// TIA Portal project "RRI" (V15.1) (continued)
   PartManagmenent.PartRecept.NazivniPodatki.CILINDRI.MOTOR4[19] := FALSE;
   PartManagmenent.PartRecept.NazivniPodatki.CILINDRI.MOTOR4[20] := FALSE;
   PartManagmenent.PartRecept.NazivniPodatki.CILINDRI.MOTOR5[1] := FALSE;
   PartManagmenent.PartRecept.NazivniPodatki.CILINDRI.MOTOR5[2] := FALSE;
   PartManagmenent.PartRecept.NazivniPodatki.CILINDRI.MOTOR5[3] := FALSE;
   PartManagmenent.PartRecept.NazivniPodatki.CILINDRI.MOTOR5[4] := FALSE;
   PartManagmenent.PartRecept.NazivniPodatki.CILINDRI.MOTOR5[5] := FALSE;
   PartManagmenent.PartRecept.NazivniPodatki.CILINDRI.MOTOR5[6] := FALSE;
   PartManagmenent.PartRecept.NazivniPodatki.CILINDRI.MOTOR5[7] := FALSE;
   PartManagmenent.PartRecept.NazivniPodatki.CILINDRI.MOTOR5[8] := FALSE;
   PartManagmenent.PartRecept.NazivniPodatki.CILINDRI.MOTOR5[9] := FALSE;
   PartManagmenent.PartRecept.NazivniPodatki.CILINDRI.MOTOR5[10] := FALSE;
   PartManagmenent.PartRecept.NazivniPodatki.CILINDRI.MOTOR5[11] := FALSE;
   PartManagmenent.PartRecept.NazivniPodatki.CILINDRI.MOTOR5[12] := FALSE;
   PartManagmenent.PartRecept.NazivniPodatki.CILINDRI.MOTOR5[13] := FALSE;
   PartManagmenent.PartRecept.NazivniPodatki.CILINDRI.MOTOR5[14] := FALSE;
   PartManagmenent.PartRecept.NazivniPodatki.CILINDRI.MOTOR5[15] := FALSE;
   PartManagmenent.PartRecept.NazivniPodatki.CILINDRI.MOTOR5[16] := FALSE;
   PartManagmenent.PartRecept.NazivniPodatki.CILINDRI.MOTOR5[17] := FALSE;
   PartManagmenent.PartRecept.NazivniPodatki.CILINDRI.MOTOR5[18] := FALSE;
   PartManagmenent.PartRecept.NazivniPodatki.CILINDRI.MOTOR5[19] := FALSE;
   PartManagmenent.PartRecept.NazivniPodatki.CILINDRI.MOTOR5[20] := FALSE;
   PartManagmenent.PartRecept.NazivniPodatki.CILINDRI.MOTOR6[1] := FALSE;
   PartManagmenent.PartRecept.NazivniPodatki.CILINDRI.MOTOR6[2] := FALSE;
   PartManagmenent.PartRecept.NazivniPodatki.CILINDRI.MOTOR6[3] := FALSE;
   PartManagmenent.PartRecept.NazivniPodatki.CILINDRI.MOTOR6[4] := FALSE;
   PartManagmenent.PartRecept.NazivniPodatki.CILINDRI.MOTOR6[5] := FALSE;
   PartManagmenent.PartRecept.NazivniPodatki.CILINDRI.MOTOR6[6] := FALSE;
   PartManagmenent.PartRecept.NazivniPodatki.CILINDRI.MOTOR6[7] := FALSE;
   PartManagmenent.PartRecept.NazivniPodatki.CILINDRI.MOTOR6[8] := FALSE;
   PartManagmenent.PartRecept.NazivniPodatki.CILINDRI.MOTOR6[9] := FALSE;
   PartManagmenent.PartRecept.NazivniPodatki.CILINDRI.MOTOR6[10] := FALSE;
   PartManagmenent.PartRecept.NazivniPodatki.CILINDRI.MOTOR6[11] := FALSE;
   PartManagmenent.PartRecept.NazivniPodatki.CILINDRI.MOTOR6[12] := FALSE;
   PartManagmenent.PartRecept.NazivniPodatki.CILINDRI.MOTOR6[13] := FALSE;
   PartManagmenent.PartRecept.NazivniPodatki.CILINDRI.MOTOR6[14] := FALSE;
   PartManagmenent.PartRecept.NazivniPodatki.CILINDRI.MOTOR6[15] := FALSE;
   PartManagmenent.PartRecept.NazivniPodatki.CILINDRI.MOTOR6[16] := FALSE;
   PartManagmenent.PartRecept.NazivniPodatki.CILINDRI.MOTOR6[17] := FALSE;
   PartManagmenent.PartRecept.NazivniPodatki.CILINDRI.MOTOR6[18] := FALSE;
   PartManagmenent.PartRecept.NazivniPodatki.CILINDRI.MOTOR6[19] := FALSE;
   PartManagmenent.PartRecept.NazivniPodatki.CILINDRI.MOTOR6[20] := FALSE;
   PartManagmenent.PartRecept.TrenutniPodatki.trenutni_pomik := 0;
   PartManagmenent.PartRecept.Oblika.s1[0] := FALSE;
   PartManagmenent.PartRecept.Oblika.s1[1] := FALSE;
   PartManagmenent.PartRecept.Oblika.s1[2] := FALSE;
   PartManagmenent.PartRecept.Oblika.s1[3] := FALSE;
   PartManagmenent.PartRecept.Oblika.s1[4] := FALSE;
   PartManagmenent.PartRecept.Oblika.s1[5] := FALSE;
   PartManagmenent.PartRecept.Oblika.s1[6] := FALSE;
   PartManagmenent.PartRecept.Oblika.s1[7] := FALSE;
   PartManagmenent.PartRecept.Oblika.s1[8] := FALSE;
   PartManagmenent.PartRecept.Oblika.s1[9] := FALSE;
   PartManagmenent.PartRecept.Oblika.s1[10] := FALSE;
   PartManagmenent.PartRecept.Oblika.s1[11] := FALSE;
   PartManagmenent.PartRecept.Oblika.s1[12] := FALSE;
   PartManagmenent.PartRecept.Oblika.s1[13] := FALSE;
   PartManagmenent.PartRecept.Oblika.s1[14] := FALSE;
   PartManagmenent.PartRecept.Oblika.s1[15] := FALSE;
   PartManagmenent.PartRecept.Oblika.s1[16] := FALSE;
   PartManagmenent.PartRecept.Oblika.s1[17] := FALSE;
   PartManagmenent.PartRecept.Oblika.s1[18] := FALSE;
   PartManagmenent.PartRecept.Oblika.s1[19] := FALSE;
   PartManagmenent.PartRecept.Oblika.s1[20] := FALSE;
   PartManagmenent.PartRecept.Oblika.s2[0] := FALSE;
   PartManagmenent.PartRecept.Oblika.s2[1] := FALSE;
   PartManagmenent.PartRecept.Oblika.s2[2] := FALSE;
   PartManagmenent.PartRecept.Oblika.s2[3] := FALSE;
   PartManagmenent.PartRecept.Oblika.s2[4] := FALSE;
   PartManagmenent.PartRecept.Oblika.s2[5] := FALSE;
   PartManagmenent.PartRecept.Oblika.s2[6] := FALSE;
   PartManagmenent.PartRecept.Oblika.s2[7] := FALSE;
   PartManagmenent.PartRecept.Oblika.s2[8] := FALSE;
   PartManagmenent.PartRecept.Oblika.s2[9] := FALSE;
   PartManagmenent.PartRecept.Oblika.s2[10] := FALSE;
   PartManagmenent.PartRecept.Oblika.s2[11] := FALSE;
   PartManagmenent.PartRecept.Oblika.s2[12] := FALSE;
   PartManagmenent.PartRecept.Oblika.s2[13] := FALSE;
   PartManagmenent.PartRecept.Oblika.s2[14] := FALSE;
   PartManagmenent.PartRecept.Oblika.s2[15] := FALSE;
   PartManagmenent.PartRecept.Oblika.s2[16] := FALSE;
   PartManagmenent.PartRecept.Oblika.s2[17] := FALSE;
   PartManagmenent.PartRecept.Oblika.s2[18] := FALSE;
   PartManagmenent.PartRecept.Oblika.s2[19] := FALSE;
   PartManagmenent.PartRecept.Oblika.s2[20] := FALSE;
   PartManagmenent.xMerkers[0] := FALSE;
   PartManagmenent.xMerkers[1] := FALSE;
END_DATA_BLOCK

DATA_BLOCK "FB_TcConvert_DB_TC1_ToolTemeprature"   // DB4
{ S7_Optimized_Access := 'TRUE' }
VERSION : 0.1
// stored: InstanceOfName FB_TcConvert
"FB_TcConvert"
BEGIN
END_DATA_BLOCK

DATA_BLOCK "FB_TcConvert_DB_TC2_ToolTemeprature"   // DB5
{ S7_Optimized_Access := 'TRUE' }
VERSION : 0.1
// stored: InstanceOfName FB_TcConvert
"FB_TcConvert"
BEGIN
END_DATA_BLOCK

DATA_BLOCK "FB_AKDstartup_DB_AKD1"   // DB6
{ S7_Optimized_Access := 'TRUE' }
VERSION : 0.1
// stored: InstanceOfName FB_AKDstartup
"FB_AKDstartup"
BEGIN
END_DATA_BLOCK

DATA_BLOCK "FB_AKDstartup_DB_TC4"   // DB7
{ S7_Optimized_Access := 'TRUE' }
VERSION : 0.1
// stored: InstanceOfName FB_AKDstartup
"FB_AKDstartup"
BEGIN
END_DATA_BLOCK

DATA_BLOCK "FB_TcConvert_DB_tc4"   // DB8
{ S7_Optimized_Access := 'TRUE' }
VERSION : 0.1
// stored: InstanceOfName FB_TcConvert
"FB_TcConvert"
BEGIN
END_DATA_BLOCK

DATA_BLOCK "FB_RTDConvert_DB_RTD1"   // DB9
{ S7_Optimized_Access := 'TRUE' }
VERSION : 0.1
// stored: InstanceOfName FB_RTDConvert
"FB_RTDConvert"
BEGIN
END_DATA_BLOCK

DATA_BLOCK "FB_RTDConvert_DB_RTD2"   // DB10
{ S7_Optimized_Access := 'TRUE' }
VERSION : 0.1
// stored: InstanceOfName FB_RTDConvert
"FB_RTDConvert"
BEGIN
END_DATA_BLOCK

DATA_BLOCK "FB_RTDConvert_DB_RTD3"   // DB11
{ S7_Optimized_Access := 'TRUE' }
VERSION : 0.1
// stored: InstanceOfName FB_RTDConvert
"FB_RTDConvert"
BEGIN
END_DATA_BLOCK

DATA_BLOCK "FB_RTDConvert_DB_RTD4"   // DB12
{ S7_Optimized_Access := 'TRUE' }
VERSION : 0.1
// stored: InstanceOfName FB_RTDConvert
"FB_RTDConvert"
BEGIN
END_DATA_BLOCK

DATA_BLOCK "LMqtt_Publisher_DB"   // DB13
{ S7_Optimized_Access := 'TRUE' }
VERSION : 0.1
// stored: InstanceOfName LMqtt_Publisher
"LMqtt_Publisher"
BEGIN
END_DATA_BLOCK

DATA_BLOCK "FB_concatScrings_DB"   // DB18
{ S7_Optimized_Access := 'TRUE' }
VERSION : 0.1
// stored: InstanceOfName FB_concatScrings
"FB_concatScrings"
BEGIN
END_DATA_BLOCK

DATA_BLOCK "DB_rPMCalculator"   // DB19
{ S7_Optimized_Access := 'TRUE' }
VERSION : 0.1
   VAR RETAIN
      Press_one : Struct
         p_trig : Bool;
         iCurrentCounter : Int;
         rCurrentSpeed : Int;
         PulseTimer : TON_TIME;
         xcalculateRPM : Bool;
      END_STRUCT;
   END_VAR
BEGIN
END_DATA_BLOCK

DATA_BLOCK "LMqtt_Publisher_DB1"   // DB22
{ S7_Optimized_Access := 'TRUE' }
VERSION : 0.1
// stored: InstanceOfName LMqtt_Publisher
"LMqtt_Publisher"
BEGIN
END_DATA_BLOCK

DATA_BLOCK "FB_concatScrings_DB1"   // DB23
{ S7_Optimized_Access := 'TRUE' }
VERSION : 0.1
// stored: InstanceOfName FB_concatScrings
"FB_concatScrings"
BEGIN
END_DATA_BLOCK

DATA_BLOCK "FB_CONCAT_STRINGS_FOR_MQTT_DB"   // DB24
{ S7_Optimized_Access := 'TRUE' }
VERSION : 0.1
// stored: InstanceOfName FB_CONCAT_STRINGS_FOR_MQTT
"FB_CONCAT_STRINGS_FOR_MQTT"
BEGIN
END_DATA_BLOCK

DATA_BLOCK "LMqtt_Publisher_1_DB"   // DB25
{ S7_Optimized_Access := 'TRUE' }
VERSION : 0.1
// stored: InstanceOfName LMqtt_Publisher_1
"LMqtt_Publisher_1"
BEGIN
END_DATA_BLOCK

DATA_BLOCK "DB_TESTWSTRING"   // DB26
{ S7_Optimized_Access := 'TRUE' }
VERSION : 0.1
   VAR
      wstring_test : WString[1000];
   END_VAR
BEGIN
END_DATA_BLOCK

DATA_BLOCK "FB_CONCAT_STRINGS_FOR_MQTT_DB_1"   // DB27
{ S7_Optimized_Access := 'TRUE' }
VERSION : 0.1
// stored: InstanceOfName FB_CONCAT_STRINGS_FOR_MQTT
"FB_CONCAT_STRINGS_FOR_MQTT"
BEGIN
END_DATA_BLOCK

DATA_BLOCK "FB_CONCAT_STRINGS_FOR_MQTT_1_DB"   // DB28
{ S7_Optimized_Access := 'TRUE' }
VERSION : 0.1
// stored: InstanceOfName FB_CONCAT_STRINGS_FOR_MQTT_1
"FB_CONCAT_STRINGS_FOR_MQTT_1"
BEGIN
END_DATA_BLOCK

DATA_BLOCK "FB_saveConcat_DB"   // DB29
{ S7_Optimized_Access := 'TRUE' }
VERSION : 0.1
// stored: InstanceOfName FB_saveConcat
"FB_saveConcat"
BEGIN
END_DATA_BLOCK

DATA_BLOCK "FB_AKD_DB_AKD1"   // DB30
{ S7_Optimized_Access := 'TRUE' }
VERSION : 0.1
// stored: InstanceOfName FB_AKD
"FB_AKD"
BEGIN
END_DATA_BLOCK

DATA_BLOCK "_AKD1"   // DB32
{ S7_Optimized_Access := 'TRUE' }
VERSION : 0.1
// stored: InstanceOfName PTC_1000_resistanceCalculation
"PTC_1000_resistanceCalculation"
BEGIN
END_DATA_BLOCK

DATA_BLOCK "FB_EgasiMotorControl_DB_M1"   // DB35
{ S7_Optimized_Access := 'TRUE' }
VERSION : 0.1
// stored: InstanceOfName FB_EgasiMotorControl
"FB_EgasiMotorControl"
BEGIN
END_DATA_BLOCK

DATA_BLOCK "DB_safetyActuator"   // DB36
{ S7_Optimized_Access := 'TRUE' }
VERSION : 0.1
   VAR RETAIN
      On_timer : Array[0..1] of TON_TIME;
      timerOut : Bool;
   END_VAR
BEGIN
END_DATA_BLOCK

DATA_BLOCK "FB_EgasiMotorControl_DB_M2"   // DB37
{ S7_Optimized_Access := 'TRUE' }
VERSION : 0.1
// stored: InstanceOfName FB_EgasiMotorControl
"FB_EgasiMotorControl"
BEGIN
END_DATA_BLOCK

DATA_BLOCK "FB_EgasiMotorControl_DB_M3"   // DB38
{ S7_Optimized_Access := 'TRUE' }
VERSION : 0.1
// stored: InstanceOfName FB_EgasiMotorControl
"FB_EgasiMotorControl"
BEGIN
END_DATA_BLOCK

DATA_BLOCK "FB_EgasiMotorControl_DB_M4"   // DB39
{ S7_Optimized_Access := 'TRUE' }
VERSION : 0.1
// stored: InstanceOfName FB_EgasiMotorControl
"FB_EgasiMotorControl"
BEGIN
END_DATA_BLOCK

DATA_BLOCK "FB_EgasiMotorControl_DB_M5"   // DB40
{ S7_Optimized_Access := 'TRUE' }
VERSION : 0.1
// stored: InstanceOfName FB_EgasiMotorControl
"FB_EgasiMotorControl"
BEGIN
END_DATA_BLOCK

DATA_BLOCK "DB_EGASI_MOTOR_BASE"   // DB41
{ S7_Optimized_Access := 'TRUE' }
VERSION : 0.1
   VAR RETAIN
      MOTOR : Array[1..5] of "EGASI_MOTOR_CONTROL";
   END_VAR
BEGIN
END_DATA_BLOCK

DATA_BLOCK "DB_PARTS_DATABASE"   // DB42
{ S7_Optimized_Access := 'TRUE' }
VERSION : 0.1
BEGIN
END_DATA_BLOCK

DATA_BLOCK "DB_RRI_Izdelki"   // DB43
{ S7_Optimized_Access := 'TRUE' }
VERSION : 0.1
   VAR RETAIN
      "1x2-Cell" : "RRI_izdelki";
      "1x4-Cell" : "RRI_izdelki";
      "1x6-Cell" : "RRI_izdelki";
      "1x8-Cell" : "RRI_izdelki";
      "2x2-Cell" : "RRI_izdelki";
      "2x4-Cell" : "RRI_izdelki";
      "2x6-Cell" : "RRI_izdelki";
      "2x8-Cell" : "RRI_izdelki";
      "39900-8" : "RRI_izdelki";
      "39900-9" : "RRI_izdelki";
   END_VAR
BEGIN
   "1x2-Cell".NazivniPodatki.st_pomikov := 2;
   "1x2-Cell".NazivniPodatki.st_celic := 2;
   "1x2-Cell".NazivniPodatki.st_vrst := 1;
   "1x4-Cell".NazivniPodatki.st_pomikov := 4;
   "1x4-Cell".NazivniPodatki.st_celic := 4;
   "1x4-Cell".NazivniPodatki.st_vrst := 1;
   "1x6-Cell".NazivniPodatki.st_pomikov := 6;
   "1x6-Cell".NazivniPodatki.st_celic := 6;
   "1x6-Cell".NazivniPodatki.st_vrst := 1;
   "1x8-Cell".NazivniPodatki.st_celic := 8;
   "1x8-Cell".NazivniPodatki.st_pomikov := 8;
   "1x8-Cell".NazivniPodatki.st_vrst := 1;
   "2x2-Cell".NazivniPodatki.st_pomikov := 2;
   "2x2-Cell".NazivniPodatki.st_celic := 2;
   "2x2-Cell".NazivniPodatki.st_vrst := 2;
   "2x4-Cell".NazivniPodatki.st_pomikov := 4;
   "2x4-Cell".NazivniPodatki.st_celic := 4;
   "2x4-Cell".NazivniPodatki.st_vrst := 2;
   "2x6-Cell".NazivniPodatki.st_pomikov := 6;
   "2x6-Cell".NazivniPodatki.st_celic := 6;
   "2x6-Cell".NazivniPodatki.st_vrst := 2;
   "2x8-Cell".NazivniPodatki.st_pomikov := 8;
   "2x8-Cell".NazivniPodatki.st_celic := 8;
   "2x8-Cell".NazivniPodatki.st_vrst := 2;
END_DATA_BLOCK

DATA_BLOCK "FB_CYLINDER_CONTROL_DB"   // DB44
{ S7_Optimized_Access := 'TRUE' }
VERSION : 0.1
// stored: InstanceOfName FB_CYLINDER_CONTROL
"FB_CYLINDER_CONTROL"
BEGIN
END_DATA_BLOCK

DATA_BLOCK "FB_VerifyTheFormLerning_DB"   // DB47
{ S7_Optimized_Access := 'TRUE' }
VERSION : 0.1
// stored: InstanceOfName FB_VerifyTheFormLerning
"FB_VerifyTheFormLerning"
BEGIN
END_DATA_BLOCK

DATA_BLOCK "DB_newGlobalDataForChangeParrt"   // DB48
{ S7_Optimized_Access := 'TRUE' }
VERSION : 0.1
   VAR RETAIN
      ud_GlobalFeedCounter : UDInt;
      DATA : "M_position";
      changePartCounter : UDInt;
      strip : Array[0..20] of "STRIP_SEGMENT";
   END_VAR
BEGIN
   DATA.POSITION_INSIDE_TOOL.M1 := 5;
   DATA.POSITION_INSIDE_TOOL.M2 := 8;
   DATA.POSITION_INSIDE_TOOL.M3 := 10;
   DATA.POSITION_INSIDE_TOOL.M4 := 14;
   DATA.POSITION_INSIDE_TOOL.M5 := 17;
   DATA.POSITION_INSIDE_TOOL.TOOL_MAX_FEED := 17;
END_DATA_BLOCK

DATA_BLOCK "FB_CYLINDER_CONTROL_PIPILINE_DB"   // DB49
{ S7_Optimized_Access := 'TRUE' }
VERSION : 0.1
// stored: InstanceOfName FB_CYLINDER_CONTROL_PIPILINE
"FB_CYLINDER_CONTROL_PIPILINE"
BEGIN
END_DATA_BLOCK

// folder: AKD

DATA_BLOCK "DB_AKD"   // DB31
{ S7_Optimized_Access := 'TRUE' }
VERSION : 0.1
BEGIN
END_DATA_BLOCK

// folder: AKD/PNU

DATA_BLOCK "AKD_PNU_DATA"   // DB33
{ S7_Optimized_Access := 'TRUE' }
VERSION : 0.1
   VAR
      AKD1 : Struct
         PNU_DATA : "PNU_DATA";
         PNU_userSETTINGS : Struct
            xRadAKDTemp : Bool;
            xReadAkdTempInC : Bool;
            PNU_const : Struct
               AKD_TEMP : Struct
                  PNU_number : Int := 2257;
                  PNU_subIndex : Int := 0;
                  PNU_type : Word := 16#43;
               END_STRUCT;
               AKD_TEMP_C : Struct
                  PNU_number : Int := 2258;
                  PNU_subIndex : Int := 0;
                  PNU_type : Word := 16#43;
               END_STRUCT;
            END_STRUCT;
         END_STRUCT;
      END_STRUCT;
   END_VAR
BEGIN
END_DATA_BLOCK

DATA_BLOCK "AKD1_PNU"   // DB34
{ S7_Optimized_Access := 'FALSE' }
AUTHOR : jcoleman
FAMILY : PNU
VERSION : 2.0
// stored: InstanceOfName AKD_PNU_v02
"AKD_PNU_v02"
BEGIN
END_DATA_BLOCK

// folder: MQTT

DATA_BLOCK "LMqtt_Status"   // DB14
{ S7_Optimized_Access := 'TRUE' }
VERSION : 0.1
   VAR
      mqtt_1 : Struct
         xtcpEsablished : Bool;   // True if the TCP connection has been
         xmqttEstavlished : Bool;   // True if the MQTT connection has been established
         xpublished : Bool;   // True, if the message has arrived successfully at
         xbusy : Bool;   // True, while a message or ping is sent to the
         xerror : Bool;   // True if there is an error
         istatusID : Int;   // State that cause the error
         status : DWord;   // Error message
      END_STRUCT;
   END_VAR
BEGIN
END_DATA_BLOCK

DATA_BLOCK "instPublisherDB"   // DB15
{ S7_Optimized_Access := 'TRUE' }
VERSION : 0.1
// stored: InstanceOfName LMqtt_Publisher
"LMqtt_Publisher"
BEGIN
END_DATA_BLOCK

DATA_BLOCK "LMqtt_Data"   // DB16
{ S7_Optimized_Access := 'TRUE' }
VERSION : 0.1
   VAR
      dataTcp : "typeTcpConnParam";
      dataMqtt : "typeMqttParam";
   END_VAR
BEGIN
   dataMqtt.connectFlag.cleanSession := 1;
   dataMqtt.connectFlag.will := 0;
   dataMqtt.connectFlag.willQoS_1 := 0;
   dataMqtt.connectFlag.willRetain := 0;
   dataMqtt.clientIdentifier := 'S7-1200-PLC';
   dataMqtt.willTopic := '/final';
   dataMqtt.willMessage := 'Das wars';
   dataTcp.hwIdentifier := 64;
   dataTcp.connectionID := 16#2;
   dataTcp.ipAdressBroker[0] := 192;
   dataMqtt.topic := 'data/s71200';
   dataMqtt.message := 'My first message';
   dataMqtt.publishFlag.qualityOfService := 1;
   dataMqtt.keepAlive := 0;
   dataTcp.localPort := 2000;
   dataTcp.mqttPort := 1883;
   dataMqtt.connectFlag.password := 0;
   dataMqtt.connectFlag.userName := 0;
   dataMqtt.userName := 'simatic';
   dataMqtt.password := 'Anna';
   dataTcp.ipAdressBroker[1] := 168;
   dataTcp.ipAdressBroker[2] := 1;
   dataTcp.ipAdressBroker[3] := 1;
END_DATA_BLOCK

DATA_BLOCK "LMqtt_publish"   // DB17
{ S7_Optimized_Access := 'TRUE' }
VERSION : 0.1
   VAR
      LMqtt : Struct
         xenable : Bool;
         epublish : Bool;
         sStringToPublish : String;
      END_STRUCT;
      randomstrinmg : String;
   END_VAR
BEGIN
END_DATA_BLOCK

// folder: MQTT/userData

DATA_BLOCK "MQTT_DB"   // DB21
{ S7_Optimized_Access := 'TRUE' }
VERSION : 0.1
   VAR RETAIN
      MQTT_CLIEENTS : Array[0..1] of "typeMqttData";
   END_VAR
   VAR
      MQTT_CLIENTS_WSTRING : Array[0..1] of "typeMqttData_1";
   END_VAR
BEGIN
   MQTT_CLIEENTS[0].mqttTcpParam.hwIdentifier := 64;
   MQTT_CLIEENTS[0].mqttTcpParam.connectionID := 16#0003;
   MQTT_CLIEENTS[0].mqttTcpParam.ipAdressBroker[0] := 16#C0;
   MQTT_CLIEENTS[0].mqttTcpParam.ipAdressBroker[1] := 16#A8;
   MQTT_CLIEENTS[0].mqttTcpParam.ipAdressBroker[2] := 16#01;
   MQTT_CLIEENTS[0].mqttTcpParam.ipAdressBroker[3] := 16#01;
   MQTT_CLIEENTS[0].mqttTcpParam.localPort := 2001;
   MQTT_CLIEENTS[0].mqttTcpParam.mqttPort := 1883;
   MQTT_CLIEENTS[0].mqttParam.connectFlag.cleanSession := TRUE;
   MQTT_CLIEENTS[0].mqttParam.clientIdentifier := 'S7-1200-PLC2';
   MQTT_CLIEENTS[0].mqttParam.willTopic := '/final2';
   MQTT_CLIEENTS[0].mqttParam.topic := 'data/s71200/RTDvalues';
   MQTT_CLIEENTS[0].mqttParam.message := '{"temperature1":                  -1.0000,"temperature2":                  -1.0000,"temperature3":                  22.8000,"temperature4":                  -1.0000}';
   MQTT_CLIEENTS[0].mqttParam.connectFlag.will := FALSE;
   MQTT_CLIEENTS[0].mqttParam.connectFlag.willQoS_1 := FALSE;
   MQTT_CLIEENTS[0].mqttParam.connectFlag.willQoS_2 := FALSE;
   MQTT_CLIEENTS[0].mqttParam.connectFlag.willRetain := FALSE;
   MQTT_CLIEENTS[0].mqttParam.connectFlag.password := FALSE;
   MQTT_CLIEENTS[0].mqttParam.connectFlag.userName := FALSE;
   MQTT_CLIEENTS[0].mqttParam.publishFlag.qualityOfService := 0;
   MQTT_CLIEENTS[0].mqttParam.publishFlag.retain := FALSE;
   MQTT_CLIEENTS[0].mqttParam.keepAlive := 16#000A;
   MQTT_CLIEENTS[0].mqttParam.packetIdentifier := 16#0010;
   MQTT_CLIEENTS[0].mqttParam.willMessage := 'das';
   MQTT_CLIEENTS[0].mqttParam.userName := 'Simatic';
   MQTT_CLIEENTS[0].mqttParam.password := 'Anna';
   MQTT_CLIEENTS[0].mqttUserControl.xEnable := TRUE;
   MQTT_CLIEENTS[0].mqttUserControl.xPusblish := FALSE;
   MQTT_CLIEENTS[0].mqttUserControl.sStringToPublish := '{"temperature1":                  -1.0000,"temperature2":                  -1.0000,"temperature3":                  22.8000,"temperature4":                  -1.0000}';
   MQTT_CLIEENTS[0].mqttUserControl.Status.xtcpEsablished := TRUE;
   MQTT_CLIEENTS[0].mqttUserControl.Status.xmqttEstavlished := TRUE;
   MQTT_CLIEENTS[0].mqttUserControl.Status.xpublished := FALSE;
   MQTT_CLIEENTS[0].mqttUserControl.Status.xbusy := FALSE;
   MQTT_CLIEENTS[0].mqttUserControl.Status.xerror := FALSE;
   MQTT_CLIEENTS[0].mqttUserControl.Status.istatusID := 0;
   MQTT_CLIEENTS[0].mqttUserControl.Status.status := 16#0000_0000;
   MQTT_CLIEENTS[1].mqttTcpParam.hwIdentifier := 0;
   MQTT_CLIEENTS[1].mqttTcpParam.connectionID := 16#0000;
   MQTT_CLIEENTS[1].mqttTcpParam.ipAdressBroker[0] := 16#00;
   MQTT_CLIEENTS[1].mqttTcpParam.ipAdressBroker[1] := 16#00;
   MQTT_CLIEENTS[1].mqttTcpParam.ipAdressBroker[2] := 16#00;
   MQTT_CLIEENTS[1].mqttTcpParam.ipAdressBroker[3] := 16#00;
   MQTT_CLIEENTS[1].mqttTcpParam.localPort := 0;
   MQTT_CLIEENTS[1].mqttTcpParam.mqttPort := 0;
   MQTT_CLIEENTS[1].mqttParam.connectFlag.cleanSession := FALSE;
   MQTT_CLIEENTS[1].mqttParam.connectFlag.will := FALSE;
   MQTT_CLIEENTS[1].mqttParam.connectFlag.willQoS_1 := FALSE;
   MQTT_CLIEENTS[1].mqttParam.connectFlag.willQoS_2 := FALSE;
   MQTT_CLIEENTS[1].mqttParam.connectFlag.willRetain := FALSE;
   MQTT_CLIEENTS[1].mqttParam.connectFlag.password := FALSE;
   MQTT_CLIEENTS[1].mqttParam.connectFlag.userName := FALSE;
   MQTT_CLIEENTS[1].mqttParam.publishFlag.qualityOfService := 0;
   MQTT_CLIEENTS[1].mqttParam.publishFlag.retain := FALSE;
   MQTT_CLIEENTS[1].mqttParam.keepAlive := 16#000A;
   MQTT_CLIEENTS[1].mqttParam.packetIdentifier := 16#0010;
   MQTT_CLIEENTS[1].mqttParam.clientIdentifier := '';
   MQTT_CLIEENTS[1].mqttParam.willTopic := '';
   MQTT_CLIEENTS[1].mqttParam.willMessage := '';
   MQTT_CLIEENTS[1].mqttParam.userName := '';
   MQTT_CLIEENTS[1].mqttParam.password := '';
   MQTT_CLIEENTS[1].mqttParam.topic := '';
   MQTT_CLIEENTS[1].mqttParam.message := '';
   MQTT_CLIEENTS[1].mqttUserControl.xEnable := FALSE;
   MQTT_CLIEENTS[1].mqttUserControl.xPusblish := FALSE;
   MQTT_CLIEENTS[1].mqttUserControl.sStringToPublish := '';
   MQTT_CLIEENTS[1].mqttUserControl.Status.xtcpEsablished := FALSE;
   MQTT_CLIEENTS[1].mqttUserControl.Status.xmqttEstavlished := FALSE;
   MQTT_CLIEENTS[1].mqttUserControl.Status.xpublished := FALSE;
   MQTT_CLIEENTS[1].mqttUserControl.Status.xbusy := FALSE;
   MQTT_CLIEENTS[1].mqttUserControl.Status.xerror := FALSE;
   MQTT_CLIEENTS[1].mqttUserControl.Status.istatusID := 0;
   MQTT_CLIEENTS[1].mqttUserControl.Status.status := 16#0000_0000;
   MQTT_CLIENTS_WSTRING[0].mqttParam.topic := 'data/s71200/testValues';
   MQTT_CLIENTS_WSTRING[0].mqttParam.password := 'Anna';
   MQTT_CLIENTS_WSTRING[0].mqttParam.userName := 'Simatic';
   MQTT_CLIENTS_WSTRING[0].mqttParam.willMessage := 'das';
   MQTT_CLIENTS_WSTRING[0].mqttParam.willTopic := '/final2';
   MQTT_CLIENTS_WSTRING[0].mqttParam.clientIdentifier := 'S7-1200-WS';
   MQTT_CLIENTS_WSTRING[0].mqttParam.packetIdentifier := 16#0010;
   MQTT_CLIENTS_WSTRING[0].mqttParam.keepAlive := 16#000A;
   MQTT_CLIENTS_WSTRING[0].mqttParam.connectFlag.cleanSession := TRUE;
   MQTT_CLIENTS_WSTRING[0].mqttTcpParam.mqttPort := 1883;
   MQTT_CLIENTS_WSTRING[0].mqttTcpParam.localPort := 2003;
   MQTT_CLIENTS_WSTRING[0].mqttTcpParam.ipAdressBroker[3] := 16#01;
   MQTT_CLIENTS_WSTRING[0].mqttTcpParam.ipAdressBroker[2] := 16#01;
   MQTT_CLIENTS_WSTRING[0].mqttTcpParam.ipAdressBroker[1] := 16#A8;
   MQTT_CLIENTS_WSTRING[0].mqttTcpParam.ipAdressBroker[0] := 16#C0;
   MQTT_CLIENTS_WSTRING[0].mqttTcpParam.connectionID := 16#0006;
   MQTT_CLIENTS_WSTRING[0].mqttTcpParam.hwIdentifier := 64;
END_DATA_BLOCK

// folder: NodeRed

DATA_BLOCK "DB_DATAFORCOMMUNICATION"   // DB1
{ S7_Optimized_Access := 'FALSE' }
VERSION : 0.1
   VAR
      rTC1_ToolTemperature1 : Real;
      rTC2_ToolTemeprature2 : Real;
      rTC3_TempEnvierment : Real;
      rTC4_Temp : Real;
      iPresaHitrost : Int;
      uPresaStevec : UDInt;
      xPresaON : Int;
      r_RTD_c0 : Real;   // temp ohišja aktuatorja
      r_RTD_c1 : Real;   // ohišje orodja
      r_RTD_c2 : Real;
      r_RTD_c3 : Real;
      r_ActuatorMaxForce : Real;
      r_ActuatorMinForce : Real;
      r_EgasiTemperaturaAktuatorja : Real;
      r_M1_temperature : Real;
      r_M2_temperature : Real;
      r_M3_temperature : Real;
      r_M4_temperature : Real;
      r_M5_temperature : Real;
      r_M1_MaxForce : Real;
      r_M2_MaxForce : Real;
      r_M3_MaxForce : Real;
      r_M4_MaxForce : Real;
      r_M5_MaxForce : Real;
      i_StevecPomika : Int;
      test : Int;
      iHMIpartNumber : Int;   // Part number -> Manual
      iHmiLastPartNumber : Int;
      iOperationMode : Int;   // 0 -> MANUAL 1->AUTO
   END_VAR
BEGIN
END_DATA_BLOCK

DATA_BLOCK "DB_MotorData"   // DB45
{ S7_Optimized_Access := 'FALSE' }
VERSION : 0.1
   VAR
      M1_status : "UDT_MotorDataStatus";
      M2_status : "UDT_MotorDataStatus";
      M3_status : "UDT_MotorDataStatus";
      M4_status : "UDT_MotorDataStatus";
      M5_status : "UDT_MotorDataStatus";
   END_VAR
BEGIN
END_DATA_BLOCK

DATA_BLOCK "DB_MotorControl"   // DB46
{ S7_Optimized_Access := 'FALSE' }
VERSION : 0.1
   VAR
      HMI_M1 : "UDT_MotorControl";
      HMI_M2 : "UDT_MotorControl";
      HMI_M3 : "UDT_MotorControl";
      HMI_M4 : "UDT_MotorControl";
      HMI_M5 : "UDT_MotorControl";
      xOverRideControl : Bool;   // 1 - HMI, 0 - PLC - MOTOR STATUS , CONTRO mode HMI
      xManualMode : Bool;
      xDEMO_or_AutomaticMode : Bool;   // 0 - automatic, 1- demo
      xHMI_resetPomikna0 : Bool;
      xHMI_Manual_or_automatic_production : Bool;   // 1-MANUAL, 0-AUTOMATIC - prodution
      DTL_forProductionID : DTL;
      Static_1 : UDInt;
   END_VAR
BEGIN
END_DATA_BLOCK

// folder: System blocks/Program resources

DATA_BLOCK "xPresaOFF"   // DB20
{ S7_Optimized_Access := 'TRUE' }
AUTHOR : Simatic
FAMILY : IEC
NAME : IEC_TMR
VERSION : 1.0
// stored: InstanceOfName IEC_TIMER
"IEC_TIMER"
BEGIN
END_DATA_BLOCK

// folder: (top level)

FUNCTION_BLOCK "FB_TcConvert"   // FB1, LAD
{ S7_Optimized_Access := 'TRUE' }
VERSION : 0.1
// Convert Thermocoupler input to the °C value
   VAR_INPUT
      i_wTC_value : Word;
      i_rCalibrationFactor : Real;
   END_VAR
   VAR_OUTPUT
      q_rTemperature : Real;
   END_VAR
   VAR RETAIN
      _rConvertedValue : Real;
   END_VAR
BEGIN

REGION Network 2 (SCL)

   //Input value 254 (DEC) = 25.5°C
   //32767 - overflow or error
   IF #i_wTC_value = 32767 THEN
       #q_rTemperature := -1.0;
       RETURN;
   END_IF;

   #q_rTemperature := WORD_TO_DINT( #i_wTC_value) / 10.0-#i_rCalibrationFactor;
END_REGION
END_FUNCTION_BLOCK

FUNCTION_BLOCK "FB_AKDstartup"   // FB2, LAD
{ S7_Optimized_Access := 'TRUE' }
VERSION : 0.1
   VAR_INPUT
      i_xFaultFeedback : Bool;   // AKD drive fault - open (0) if error
      i_xStart : Bool;   // Run startup Sequence
   END_VAR
   VAR_OUTPUT
      q_xHwEnable : Bool;
      q_xSTOEnable : Bool;
      q_xAKDPower : Bool;
      q_xSoftwareEnable : Bool;
   END_VAR
   VAR
      TON_TIMER : Array[0..1] of TON_TIME;
      TOFF_TIMER : Array[0..1] of TOF_TIME;
   END_VAR
BEGIN

REGION Network 1
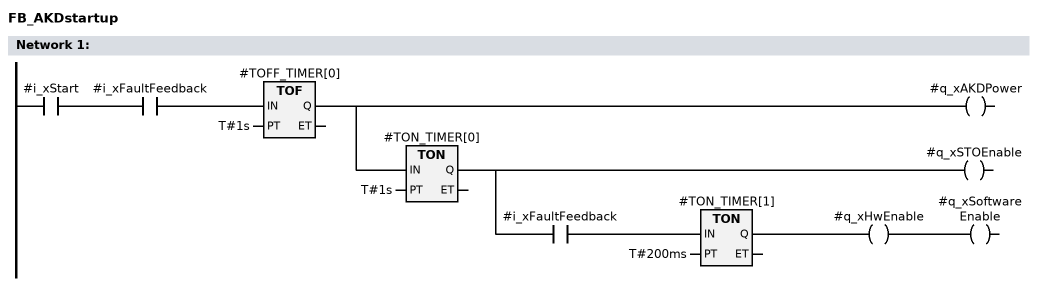
   #TOFF_TIMER[0].TOF(IN := #i_xStart AND #i_xFaultFeedback, PT := T#1s);
   #q_xAKDPower := #TOFF_TIMER[0].Q;
   #TON_TIMER[0].TON(IN := #TOFF_TIMER[0].Q, PT := T#1s);
   #q_xSTOEnable := #TON_TIMER[0].Q;
   #TON_TIMER[1].TON(IN := #TON_TIMER[0].Q AND #i_xFaultFeedback, PT := T#200ms);
   #q_xHwEnable := #TON_TIMER[1].Q;
   #q_xSoftwareEnable := #TON_TIMER[1].Q;
END_REGION
END_FUNCTION_BLOCK

FUNCTION_BLOCK "FB_RTDConvert"   // FB3, LAD
{ S7_Optimized_Access := 'TRUE' }
VERSION : 0.1
   VAR_INPUT
      i_wRTD_value : Word;
      i_rCalibrationFactor : Real;
   END_VAR
   VAR_OUTPUT
      q_rTemperature : Real;
   END_VAR
BEGIN

REGION Network 2 (SCL)

   //Input value 254 (DEC) = 25.5°C
   //32767 - overflow or error
   IF #i_wRTD_value = 32767 THEN
       #q_rTemperature := -1.0;
       RETURN;
   END_IF;

   #q_rTemperature := WORD_TO_DINT(#i_wRTD_value) / 10.000 - #i_rCalibrationFactor;
END_REGION
END_FUNCTION_BLOCK

FUNCTION_BLOCK "LMqtt_Publisher"   // FB4, SCL
{ S7_Optimized_Access := 'TRUE' }
VERSION : 0.1
   VAR_INPUT
      enable : Bool;
      publish : Bool;
      tcpConnParam : "typeTcpConnParam";
      mqttParam : "typeMqttParam";
   END_VAR
   VAR_OUTPUT
      tcpEstablished : Bool;
      mqttEstablished : Bool;
      published : Bool;
      busy : Bool;
      error : Bool;
      status : DWord;
      statusID : Int;
   END_VAR
   VAR
      statTcpConnParam : TCON_IP_v4;
      instTcpConnect : TCON;
      instTcpSend : TSEND;
      instTcpRCV : TRCV;
      instTcpDisconnect : TDISCON;
      instWatchDog : TON_TIME;
      instKeepAlive : TON_TIME;
      statStateMQTT : Int;
      statStateMQTTinternal : Int;
      statStateTCP : Int;
      statLastState : Int;
      statConnectLenght : Int;
      statCorrectOffset : Int;
      statSendLenght : Int;
      statConnectEncodedLenght : Int;
      statConnectLenghtOffset : Int;
      statKeepAliveTime : Time;
      statI : Int;
      statPacketID : Word;
      statPacketIDAck : Word;
      statRcvLen : UDInt;
      statPublishOld : Bool;
      statReConnect : Bool;
      statEnableOld : Bool;
      statMqttResetOld : Bool;
      statTriggerWatchDog : Bool;
      statTriggerKeepAlive : Bool;
      statNewDataRcv : Bool;
      statKeepAliveOff : Bool;
      statSendBuffer : Array[1..1000] of Byte;
      statRcvBuffer : Array[1..200] of Byte;
   END_VAR
   VAR_TEMP
      tempStringToChar : Array[0..255] of Char;
      tempCountChars : UInt;
      tempLenght : Word;
   END_VAR
   VAR CONSTANT
      TCP_PARAM : Int := 1;
      TCP_DISCONNECT : Int := -1;
      TCP_ERROR : Int := -2;
      TCP_CONNECTED : Int := 3;
      TCP_CONNECTING : Int := 2;
      MQTT_CONNECT_FLAG_CHECK : Int := 10;
      MQTT_CONNECT : Int := 11;
      MQTT_PUBLISH : Int := 13;
      MQTT_DISCONNECT : Int := 15;
      MQTT_CONNACK : Int := 12;
      MQTT_PUBACK : Int := 14;
      MQTT_PING : Int := 17;
      MQTT_PINGRESP : Int := 18;
      MQTT_PUBREL : Int := 19;
      MQTT_PUBCOMP : Int := 20;
      MQTT_IDLE : Int;
      MQTT_CONNECTED : Int := 16;
      MQTT_DISCONNECTED : Int := -11;
      MQTT_ERROR : Int := -12;
      IDLE : Int;
      TIME_MONITORING : Int := 20;
      WATCHDOG_TIME : Time := t#30s;
      MQTT_MSG_TYPE_CONNACK : Int := 32;
      MQTT_MSG_TYPE_DISCONNECT : Int := 224;
      MQTT_MSG_TYPE_PUBACK : Int := 64;
      MQTT_MSG_TYPE_PUBREC : Int := 80;
      MQTT_MSG_TYPE_PUBCOM : Int := 112;
      MQTT_MSG_TYPE_PING : Int := 192;
      MQTT_MSG_TYPE_PINGRESP : Int := 208;
      MQTT_CONNACK_ACCEPTED : Int;
      MQTT_PORT : Word := 16#22B3;
      MQTT_PROTOCOL_NAME : String := 'MQTT';
      MQTT_ERROR_WILL_FLAG : Word := 16#80F0;
      MQTT_ERROR_QOS_FLAG : Word := 16#80F1;
      MQTT_ERROR_PACKETID : Word := 16#80F2;
      MQTT_ERROR_KEEPALIVE : Word := 16#80F3;
   END_VAR
   // statTcpConnParam.ActiveEstablished := true;
BEGIN
   //=============================================================================
   //SIEMENES AG
   //(c)Copyright 2016 All Rights Reserved
   //-----------------------------------------------------------------------------
   //Library:       (that the source is dedicated to)
   //Tested with:   (target system with FW Version)
   //Engineering:   TIA Portal V15
   //Restrictions:  (OB types, etc.)
   //Requirements:  (hardware, technological package, memory needed, etc.)
   //Functionality: MQTT
   //-----------------------------------------------------------------------------
   //Change log table:
   //Version  Date       Expert in charge Changes applied
   //01.00.00 dd.mm.yyyy (name of expert) First released version
   //=============================================================================
   //Establish TCP Connection to be ready for MQTT

   IF #enable
       AND NOT #statEnableOld
   THEN
       #statStateTCP := #TCP_PARAM;
       #statStateMQTT := #MQTT_DISCONNECTED;
       #instWatchDog.IN := false;
       #statPublishOld := #publish;
       #error := 0;
       #status := 0;
       #statusID := 0;
   END_IF;

   IF NOT #enable
       AND #statEnableOld
   THEN
       IF #statStateTCP = #TCP_CONNECTED AND
           #statStateMQTT = #MQTT_DISCONNECTED
       THEN
           #statStateTCP := #TCP_DISCONNECT;
       END_IF;
       IF #statStateTCP = #TCP_CONNECTED AND
           #statStateMQTT <> #MQTT_DISCONNECTED
       THEN
           #statStateMQTT := #MQTT_DISCONNECT;
       END_IF;
       IF #statStateTCP = #TCP_CONNECTING
           OR  #statStateTCP = #IDLE
       THEN

           #statStateMQTT := #MQTT_DISCONNECTED;
           #statStateTCP := #IDLE;
       END_IF;
   END_IF;

    #instWatchDog(IN := #statTriggerWatchDog,PT := #WATCHDOG_TIME);

   REGION State maschine TCP
       CASE #statStateTCP OF
           #IDLE:
               IF NOT #error
               THEN
                   #status := 0;
                   #statusID := 0;

               END_IF;
               #statTcpConnParam.ID := #tcpConnParam.connectionID;
               #instTcpDisconnect(ID := #statTcpConnParam.ID);
               #instTcpConnect(ID := #statTcpConnParam.ID,
                               CONNECT := #statTcpConnParam);
               #published := 0;
               #busy := false;
               #mqttEstablished := false;
               #statMqttResetOld := 0;
               #tcpEstablished := false;
               #statStateMQTT := #MQTT_DISCONNECTED;
               #statStateMQTTinternal := #IDLE;
               #statTriggerWatchDog := false;
               #statTriggerKeepAlive := 0;
               IF #statLastState=#TCP_DISCONNECT
               THEN
                   #error := 0;
                   END_IF;
           #TCP_CONNECTED:
               ;
               //Check TCP Connection
               IF #instTcpRCV.STATUS > w#16#80C0
               THEN
                   #statStateTCP := #TCP_ERROR;
                   #statusID := #TCP_CONNECTED;
               END_IF;
               #statLastState := #TCP_CONNECTED;
           #TCP_PARAM:
               #statTcpConnParam.InterfaceId := #tcpConnParam.hwIdentifier;
               #statTcpConnParam.ID := #tcpConnParam.connectionID;
               #statTcpConnParam.LocalPort := #tcpConnParam.localPort;
               #statTcpConnParam.RemotePort := #tcpConnParam.mqttPort;
               #statTcpConnParam.ActiveEstablished := true;
               #statTcpConnParam.RemoteAddress.ADDR[1] := #tcpConnParam.ipAdressBroker[0];
               #statTcpConnParam.RemoteAddress.ADDR[2] := #tcpConnParam.ipAdressBroker[1];
               #statTcpConnParam.RemoteAddress.ADDR[3] := #tcpConnParam.ipAdressBroker[2];
               #statTcpConnParam.RemoteAddress.ADDR[4] := #tcpConnParam.ipAdressBroker[3];

             #statStateTCP := #TCP_CONNECTING;
           #TCP_CONNECTING:
               REGION TCP Connect
                   #statTriggerWatchDog := true;
                   #instTcpConnect.REQ := NOT #instTcpConnect.REQ XOR #instTcpConnect.BUSY;
                   #instTcpConnect(ID := #statTcpConnParam.ID,
                                   CONNECT := #statTcpConnParam);

                   IF (#instTcpConnect.DONE)
                       AND (#instTcpConnect.BUSY = 0)
                       AND (#instTcpConnect.REQ)
                   THEN
                       #instTcpConnect.REQ := false;
                       #tcpEstablished := true;
                       #statStateTCP := #TCP_CONNECTED;
                       #statTriggerWatchDog := false;
                   ELSIF (#instTcpConnect.ERROR)
                   THEN
                       #statusID := #TCP_CONNECTING;
                       #instTcpConnect.REQ := false;
                       #statStateTCP := #TCP_ERROR;
                   END_IF;
               END_REGION

           #TCP_DISCONNECT:
               REGION TCP Disconnect
                   #instTcpDisconnect.REQ := NOT #instTcpDisconnect.REQ XOR #instTcpDisconnect.BUSY;
                   #statTriggerWatchDog := false;
                   #instTcpDisconnect(ID := #statTcpConnParam.ID);

                   IF (#instTcpDisconnect.DONE)
                   THEN
                       //Done with success
                       #instTcpDisconnect.REQ := false;
                       #statLastState := #TCP_DISCONNECT;
                       #statStateTCP := #IDLE;
                   ELSIF (#instTcpDisconnect.ERROR)
                   THEN
                       #statusID := #TCP_DISCONNECT;
                       #instTcpDisconnect.REQ := false;
                       #statStateTCP := #TCP_ERROR;
                   END_IF;
               END_REGION
               ;
           #TCP_ERROR:
               REGION Errorhandling
                   #error := true;
                   #statStateMQTT := #MQTT_DISCONNECTED;
                   #statStateMQTTinternal := #IDLE;
                   #tcpEstablished := false;
                   #mqttEstablished := false;
                   #published := false;
                   #statTriggerWatchDog := false;
                   #instTcpConnect.REQ := false;
                       CASE #statusID OF
                           #TCP_CONNECTING:
                               #statStateTCP := #IDLE;
                               #status := #instTcpConnect.STATUS;
                           #TCP_CONNECTED:
                               #statStateTCP := #TCP_DISCONNECT;
                               #status := #instTcpRCV.STATUS;
                           #TCP_DISCONNECT:
                               //pointless for a retry at TDISCON
                               #statStateTCP := #IDLE;
                               #status := #instTcpDisconnect.STATUS;
                           #TIME_MONITORING:
                               IF (#statLastState = #TCP_CONNECTED)
                               THEN
                                   #statStateTCP := #TCP_DISCONNECT;
                                   #status := #instTcpRCV.STATUS;
                               ELSE
                                   #statStateTCP := #IDLE;
                                   #status := #instTcpConnect.STATUS;
                               END_IF;
                           ELSE
                               ;
                       END_CASE;
               END_REGION
               ;
           ELSE
               ;
       END_CASE;
   END_REGION
   #statEnableOld := #enable;
   REGION WatchDog
       IF #instWatchDog.Q = true
       THEN
           #statStateTCP := #TCP_ERROR;
           #statusID := #TIME_MONITORING;
       END_IF;
   END_REGION

   REGION OUC blocks

       #instTcpSend(ID:=#statTcpConnParam.ID,
                     DATA:=#statSendBuffer);
        #instTcpRCV(EN_R:=true,
                    ID:=#statTcpConnParam.ID,
                   LEN:=0,
                   ADHOC:=1,
                   RCVD_LEN=>#statRcvLen,
                   DATA:=#statRcvBuffer);
       IF #instTcpRCV.RCVD_LEN > 0 THEN
           #statNewDataRcv := 1;
       END_IF;

   END_REGION

   //Bring Statemachine in a definded state, if TCP Connection breaks
   IF #statStateMQTT > 0 AND
       #statStateTCP <> #TCP_CONNECTED
   THEN
       #statStateMQTT := #MQTT_DISCONNECTED;
       #instTcpSend.REQ := 0;
   END_IF;

   //MQTT makes no sense without an established TCP
   IF NOT (#statStateTCP = #TCP_CONNECTED)
   THEN
       RETURN;
   END_IF;




    #instKeepAlive(IN := #statTriggerKeepAlive,
                   PT := #statKeepAliveTime);
       CASE #statStateMQTT OF
           #MQTT_DISCONNECTED:
               #mqttEstablished := false;
               #statPublishOld := #publish;
               #statStateMQTT := #MQTT_CONNECT_FLAG_CHECK;
               #statStateMQTTinternal := #IDLE;
               #statTriggerKeepAlive := 0;
               #statKeepAliveOff := false;
               #statPacketID := #mqttParam.packetIdentifier;

           #MQTT_CONNECT_FLAG_CHECK:
               #busy := 1;
               //validate flags
               IF #mqttParam.connectFlag.willRetain
                   AND NOT #mqttParam.connectFlag.will
               THEN
                   #statStateMQTT := #MQTT_ERROR;
                   #statusID := #MQTT_CONNECT_FLAG_CHECK;
                   #status := #MQTT_ERROR_WILL_FLAG;
               ELSE
                   IF NOT #mqttParam.connectFlag.will
                       AND (#mqttParam.connectFlag.willQoS_1 OR #mqttParam.connectFlag.willQoS_2)
                   THEN
                       #statStateMQTT := #MQTT_ERROR;
                       #statusID := #MQTT_CONNECT_FLAG_CHECK;
                       #status := #MQTT_ERROR_QOS_FLAG;
                   ELSE
                       IF (#mqttParam.connectFlag.willQoS_1
                           AND #mqttParam.connectFlag.willQoS_2)
                       THEN
                           #statStateMQTT := #MQTT_ERROR;
                           #statusID := #MQTT_CONNECT_FLAG_CHECK;
                           #status := #MQTT_ERROR_QOS_FLAG;
                       ELSE;
                        #statStateMQTT := #MQTT_CONNECT;
                       END_IF;
                   END_IF;

               END_IF;
               IF (WORD_TO_INT(#mqttParam.keepAlive) = 0)
               THEN
                   #statKeepAliveOff := true;
               END_IF;
               IF (WORD_TO_INT(#mqttParam.keepAlive) < 2)
                   AND
                   (WORD_TO_INT(#mqttParam.keepAlive) > 0)
               THEN
                   #statStateMQTT := #MQTT_ERROR;
                   #statusID := #MQTT_CONNECT_FLAG_CHECK;
                   #status := #MQTT_ERROR_KEEPALIVE;
               END_IF;
               IF (WORD_TO_INT(#mqttParam.keepAlive) > 2)
               THEN
                   #statKeepAliveOff := false;
               END_IF;
           #MQTT_CONNECT:
                REGION MQTT Connect

                   //Calculate Remaining Lenght
                   #statConnectLenght := 10 + LEN(IN := #mqttParam.clientIdentifier) + 2;
                   IF #mqttParam.connectFlag.userName
                   THEN
                       #statConnectLenght := #statConnectLenght + LEN(IN := #mqttParam.userName) + 2;
                   END_IF;
                   IF #mqttParam.connectFlag.password
                   THEN
                       #statConnectLenght := #statConnectLenght + LEN(IN := #mqttParam.password) + 2;
                   END_IF;
                   IF #mqttParam.connectFlag.will
                   THEN
                       #statConnectLenght := #statConnectLenght + LEN(IN := #mqttParam.willMessage) + LEN(IN := #mqttParam.willTopic) + 4;
                   END_IF;
                   #statConnectLenghtOffset := 0;
                   //Build Telegram
                   //Fixed Header
                   #statSendBuffer[1] := 16#10;

                   #statSendLenght :=#statConnectLenght;
                   WHILE (#statConnectLenght > 0)
                   DO
                       #statConnectEncodedLenght := #statConnectLenght MOD 128;
                       #statConnectLenght := #statConnectLenght / 128;
                       // if there are more data to encode, set the top bit of this byte
                       IF #statConnectLenght > 0
                       THEN
                           #statConnectEncodedLenght := #statConnectEncodedLenght OR 128;
                           #statSendBuffer[2 + #statConnectLenghtOffset] := INT_TO_BYTE(#statConnectEncodedLenght);
                           #statConnectLenghtOffset := #statConnectLenghtOffset + 1;
                       ELSE
                           #statSendBuffer[2 + #statConnectLenghtOffset] := INT_TO_BYTE(#statConnectEncodedLenght);
                       END_IF;
                   END_WHILE;
                   #statSendLenght := #statSendLenght + #statConnectLenghtOffset;
                   //Variable Header
                   //Protocol name
                   #statSendBuffer[3 + #statConnectLenghtOffset] := 0;
                   #statSendBuffer[4 + #statConnectLenghtOffset] := 4;
                   #statSendBuffer[5 + #statConnectLenghtOffset] := 'M';
                   #statSendBuffer[6 + #statConnectLenghtOffset] := 'Q';
                   #statSendBuffer[7 + #statConnectLenghtOffset] := 'T';
                   #statSendBuffer[8 + #statConnectLenghtOffset] := 'T';
                   //Protocol Level
                   #statSendBuffer[9 + #statConnectLenghtOffset] := 4;
                   //Connect Flags
                   #statSendBuffer[10 + #statConnectLenghtOffset].%X0 := 0;
                   #statSendBuffer[10 + #statConnectLenghtOffset].%X1 := #mqttParam.connectFlag.cleanSession;
                   #statSendBuffer[10 + #statConnectLenghtOffset].%X2 := #mqttParam.connectFlag.will;
                   #statSendBuffer[10 + #statConnectLenghtOffset].%X3 := #mqttParam.connectFlag.willQoS_1;
                   #statSendBuffer[10 + #statConnectLenghtOffset].%X4 := #mqttParam.connectFlag.willQoS_2;
                   #statSendBuffer[10 + #statConnectLenghtOffset].%X5 := #mqttParam.connectFlag.willRetain;
                   #statSendBuffer[10 + #statConnectLenghtOffset].%X6 := #mqttParam.connectFlag.password;
                   #statSendBuffer[10 + #statConnectLenghtOffset].%X7 := #mqttParam.connectFlag.userName;
                   //Keep Alive in sec
                  #statSendBuffer[11 + #statConnectLenghtOffset] := #mqttParam.keepAlive.%B1;
                  #statSendBuffer[12 + #statConnectLenghtOffset] := #mqttParam.keepAlive.%B0;
                   //Payload
                   //ClientIdentifier
                   #tempLenght := INT_TO_WORD(LEN(IN := #mqttParam.clientIdentifier));
                   #statSendBuffer[13 + #statConnectLenghtOffset] := #tempLenght.%B1;
                   #statSendBuffer[14 + #statConnectLenghtOffset] := #tempLenght.%B0;
                   Strg_TO_Chars(Strg := #mqttParam.clientIdentifier,
                                 pChars := 0,
                                 Cnt => #tempCountChars,
                                 Chars := #tempStringToChar);
                   FOR #statI := 0 TO UINT_TO_INT(#tempCountChars - 1) DO
                       #statSendBuffer[15 + #statConnectLenghtOffset + #statI] := #tempStringToChar[#statI];
                   END_FOR;
                   #statConnectLenghtOffset := #statConnectLenghtOffset + #statI;
                   //WillTopic and WillMessage
                   IF #mqttParam.connectFlag.will THEN
                       #statCorrectOffset := 0;
                       #tempLenght:=INT_TO_WORD(LEN(IN := #mqttParam.willTopic));
                       #statSendBuffer[15 + #statConnectLenghtOffset] := #tempLenght.%B1;
                       #statSendBuffer[16 + #statConnectLenghtOffset] := #tempLenght.%B0;
                       Strg_TO_Chars(Strg := #mqttParam.willTopic,
                                     pChars := 0,
                                     Cnt => #tempCountChars,
                                     Chars := #tempStringToChar);
                       FOR #statI := 0 TO UINT_TO_INT(#tempCountChars - 1) DO
                           #statSendBuffer[17 + #statConnectLenghtOffset + #statI] := #tempStringToChar[#statI];
                       END_FOR;
                       #statConnectLenghtOffset := #statConnectLenghtOffset + #statI;

                       #tempLenght:=INT_TO_WORD(LEN(IN := #mqttParam.willMessage));
                       #statSendBuffer[17 + #statConnectLenghtOffset] := #tempLenght.%B1;
                       #statSendBuffer[18 + #statConnectLenghtOffset] := #tempLenght.%B0;
                       Strg_TO_Chars(Strg := #mqttParam.willMessage,
                                     pChars := 0,
                                     Cnt => #tempCountChars,
                                     Chars := #tempStringToChar);
                       FOR #statI := 0 TO UINT_TO_INT(#tempCountChars - 1) DO
                           #statSendBuffer[19 + #statConnectLenghtOffset + #statI] := #tempStringToChar[#statI];
                       END_FOR;
                       #statConnectLenghtOffset := #statConnectLenghtOffset + #statI;
                   ELSE
                       #statCorrectOffset := 4;
                   END_IF;
                   //UserName
                   IF #mqttParam.connectFlag.userName THEN
                       #tempLenght := INT_TO_WORD(LEN(IN := #mqttParam.userName));
                       #statSendBuffer[19 + #statConnectLenghtOffset - #statCorrectOffset] := #tempLenght.%B1;
                       #statSendBuffer[20 + #statConnectLenghtOffset - #statCorrectOffset] := #tempLenght.%B0;
                       Strg_TO_Chars(Strg := #mqttParam.userName,
                                     pChars := 0,
                                     Cnt => #tempCountChars,
                                     Chars := #tempStringToChar);
                       FOR #statI := 0 TO UINT_TO_INT(#tempCountChars - 1) DO
                           #statSendBuffer[21 + #statConnectLenghtOffset + #statI-#statCorrectOffset] := #tempStringToChar[#statI];
                       END_FOR;
                       #statConnectLenghtOffset := #statConnectLenghtOffset + #statI;
                   END_IF;
                   //Password
                   IF #mqttParam.connectFlag.password THEN
                       #tempLenght := INT_TO_WORD(LEN(IN := #mqttParam.password));
                       #statSendBuffer[21 + #statConnectLenghtOffset - #statCorrectOffset] := #tempLenght.%B1;
                       #statSendBuffer[22 + #statConnectLenghtOffset - #statCorrectOffset] := #tempLenght.%B0;
                       Strg_TO_Chars(Strg := #mqttParam.password,
                                     pChars := 0,
                                     Cnt => #tempCountChars,
                                     Chars := #tempStringToChar);
                       FOR #statI := 0 TO UINT_TO_INT(#tempCountChars - 1) DO
                           #statSendBuffer[23 + #statConnectLenghtOffset + #statI-#statCorrectOffset] := #tempStringToChar[#statI];
                       END_FOR;
                       #statConnectLenghtOffset := #statConnectLenghtOffset + #statI;
                   END_IF;

